
   //Convert the 3rd octet string to numerical value
   STRG_VAL(IN := #tempOctetString,
            FORMAT := W#16#0000,
            P := 1,
            OUT => #tempUInt);
   IF #tempUInt > #MAX_USINT
   THEN
     #error := TRUE;
     #status := #WRONG_VALUE_POS3;
     RETURN;
   ELSE
     #tempIpAdressTaddr.REM_IP_ADDR[3] := UINT_TO_BYTE(#tempUInt);
   END_IF;

   // Process the 4th octet of the IP Address
   #tempCharPosition := FIND(IN1 := #tempAddressString, IN2 := '.');
   IF #tempCharPosition > #NO_POS THEN
     #error := TRUE;
     #status := #WRONG_VALUE_POS4;
     RETURN;
   ELSE
     #tempCharPosition := FIND(IN1 := #tempAddressString, IN2 := ':');
   END_IF;

   // Check if Port number added
   #tempPortNumberIsSpecified := (#tempCharPosition > #NO_POS);
   IF #tempCharPosition > #MAX_CHAR_FOR_PORT_PART THEN
     #error := TRUE;
     #status := #WRONG_VALUE_PORT;
     RETURN;
   END_IF;
   IF NOT #tempPortNumberIsSpecified THEN
     #tempCharPosition := LEN(#tempAddressString) + 1;
   END_IF;

   #tempOctetString := LEFT(IN := #tempAddressString, L := #tempCharPosition - 1);
   // Check if string is empty
   IF #tempOctetString = #EMPTY_STRING THEN
     #error := TRUE;
     #status := #WRONG_VALUE_POS4;
     RETURN;
   ELSE
     #tempAddressString := DELETE(IN := #tempAddressString, P := 1, L := #tempCharPosition);
   END_IF;

   // Convert the 4th octet string to numerical value
   STRG_VAL(IN := #tempOctetString,
            FORMAT := W#16#0000,
            P := 1,
            OUT => #tempUInt);

   IF #tempUInt > #MAX_USINT THEN
     #error := TRUE;
     #status := #WRONG_VALUE_POS4;
     RETURN;
   ELSE
     #tempIpAdressTaddr.REM_IP_ADDR[4] := UINT_TO_BYTE(#tempUInt);
   END_IF;

   // If the string contains a port number too, parse it
   IF #tempPortNumberIsSpecified THEN
     // Convert the port number string to numerical value
     STRG_VAL(IN := #tempAddressString,
              FORMAT := W#16#0000,
              P := 1,
              OUT => #tempUInt);
     IF #tempUInt > #MAX_UINT OR #tempUInt = 0 THEN
       #error := TRUE;
       #status := #WRONG_VALUE_PORT;
       RETURN;
     ELSE
       #tempIpAdressTaddr.REM_PORT_NR := #tempUInt;
     END_IF;
   END_IF;

   // Write Outputs
   #LGF_StringToTaddr := #tempIpAdressTaddr;
END_FUNCTION

ORGANIZATION_BLOCK "Main"   // OB1, LAD, ProgramCycle
TITLE = "Main Program Sweep (Cycle)"
{ S7_Optimized_Access := 'TRUE' }
VERSION : 0.1
   VAR_INPUT
      Initial_Call : Bool;   // Initial call of this OB
      Remanence : Bool;   // =True, if remanent data are available
   END_VAR
   VAR_TEMP
      tmpI : Int;
      tmpI2 : Int;
   END_VAR
BEGIN

REGION Network 2
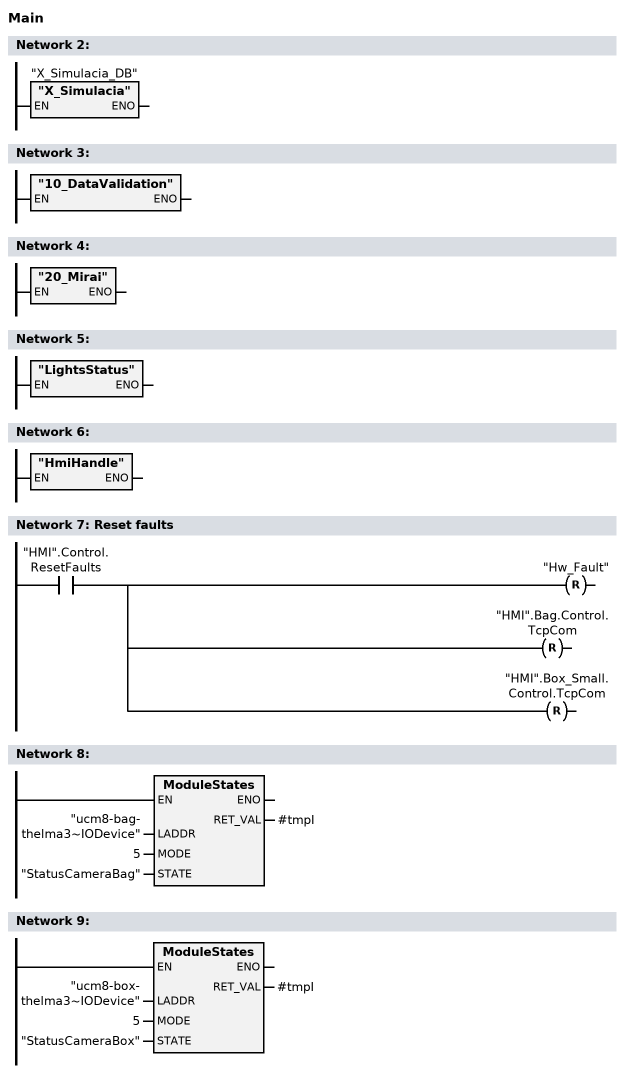
   RUNG wire#powerrail
      "X_Simulacia_DB"()
   END_RUNG
   // the same network as SCL:
   "X_Simulacia_DB"();   // "X_Simulacia"
END_REGION

REGION Network 3
   RUNG wire#powerrail
      "10_DataValidation"()
   END_RUNG
   // the same network as SCL:
   "10_DataValidation"();
END_REGION

REGION Network 4
   RUNG wire#powerrail
      "20_Mirai"()
   END_RUNG
   // the same network as SCL:
   "20_Mirai"();
END_REGION

REGION Network 5
   RUNG wire#powerrail
      "LightsStatus"()
   END_RUNG
   // the same network as SCL:
   "LightsStatus"();
END_REGION

REGION Network 6
   RUNG wire#powerrail
      "HmiHandle"()
   END_RUNG
   // the same network as SCL:
   "HmiHandle"();
END_REGION

REGION Network 7: Reset faults
   RUNG wire#powerrail
      Contact( "HMI".Control.ResetFaults )
      wire#w1
      R_Coil( "Hw_Fault" )
   END_RUNG
   RUNG wire#w1
      R_Coil( "HMI".Bag.Control.TcpCom )
   END_RUNG
   RUNG wire#w1
      R_Coil( "HMI".Box_Small.Control.TcpCom )
   END_RUNG
   // the same network as SCL:
   IF "HMI".Control.ResetFaults THEN
       "Hw_Fault" := FALSE;
       "HMI".Bag.Control.TcpCom := FALSE;
       "HMI".Box_Small.Control.TcpCom := FALSE;
   END_IF;
END_REGION

REGION Network 8
   // no SCL statement known for ModuleStates: written as a call
   #tmpI := ModuleStates(LADDR := "ucm8-bag-thelma3~IODevice", MODE := 5, STATE := "StatusCameraBag");
END_REGION

REGION Network 9
   // no SCL statement known for ModuleStates: written as a call
   #tmpI := ModuleStates(LADDR := "ucm8-box-thelma3~IODevice", MODE := 5, STATE := "StatusCameraBox");
END_REGION
END_ORGANIZATION_BLOCK

ORGANIZATION_BLOCK "Rack or station failure"   // OB86, LAD, RackStationFailure
{ S7_Optimized_Access := 'TRUE' }
VERSION : 0.1
   VAR_INPUT
      LADDR : Hw_Device;   // Hardware identifier
      Event_Class : Byte;   // Event class
      Fault_ID : Byte;   // Fault identifier
   END_VAR
BEGIN

REGION Network 1
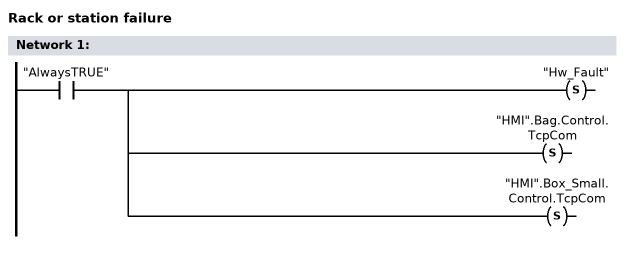
   RUNG wire#powerrail
      Contact( "AlwaysTRUE" )
      wire#w1
      S_Coil( "Hw_Fault" )
   END_RUNG
   RUNG wire#w1
      S_Coil( "HMI".Bag.Control.TcpCom )
   END_RUNG
   RUNG wire#w1
      S_Coil( "HMI".Box_Small.Control.TcpCom )
   END_RUNG
   // the same network as SCL:
   IF "AlwaysTRUE" THEN
       "Hw_Fault" := TRUE;
       "HMI".Bag.Control.TcpCom := TRUE;
       "HMI".Box_Small.Control.TcpCom := TRUE;
   END_IF;
END_REGION
END_ORGANIZATION_BLOCK

ORGANIZATION_BLOCK "Startup"   // OB100, LAD, Startup
TITLE = "Complete Restart"
{ S7_Optimized_Access := 'TRUE' }
VERSION : 0.1
   VAR_INPUT
      LostRetentive : Bool;   // True if retentive data are lost
      LostRTC : Bool;   // True if date and time are lost
   END_VAR
BEGIN

REGION Network 1
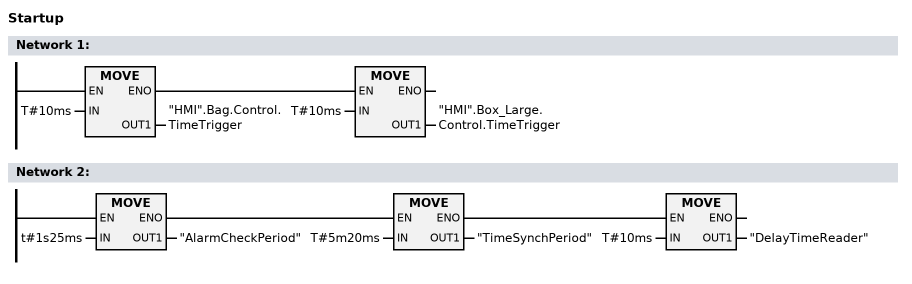
   RUNG wire#powerrail
      Move(in := T#10ms, out1 => "HMI".Bag.Control.TimeTrigger)
      Move(in := T#10ms, out1 => "HMI".Box_Large.Control.TimeTrigger)
   END_RUNG
   // the same network as SCL:
   "HMI".Bag.Control.TimeTrigger := T#10ms;
   "HMI".Box_Large.Control.TimeTrigger := T#10ms;
END_REGION

REGION Network 2
   RUNG wire#powerrail
      Move(in := t#1s25ms, out1 => "AlarmCheckPeriod")
      Move(in := T#5m20ms, out1 => "TimeSynchPeriod")
      Move(in := T#10ms, out1 => "DelayTimeReader")
   END_RUNG
   // the same network as SCL:
   "AlarmCheckPeriod" := t#1s25ms;
   "TimeSynchPeriod" := T#5m20ms;
   "DelayTimeReader" := T#10ms;
END_REGION
END_ORGANIZATION_BLOCK

ORGANIZATION_BLOCK "Programming error"   // OB121, LAD, ProgrammingError
{ S7_Optimized_Access := 'TRUE' }
VERSION : 0.1
   VAR_INPUT
      BlockNr : UInt;   // Number of causing block
      Reaction : USInt;   // 0:ignore, 1:substitute, 2:skip
      Fault_ID : Byte;   // Fault identifier
      BlockType : USInt;   // 16#01:OB, 16#02:FC, 16#03:FB, 16#04:SFC, 16#05:SFB, 16#06:DB: Type of block causing the error
      Area : USInt;   // Area where the error occured
      DBNr : DB_ANY;   // DB number if Area = DB or DI
      Csg_OBNr : OB_Any;   // Number of OB causing the error
      Csg_Prio : USInt;   // Priority of OB causing the error
      Width : USInt;   // 0:bit, 1:byte, 2:word, 3:dword, 4:lword
   END_VAR
BEGIN
END_ORGANIZATION_BLOCK

(* ===== HMI "HMI_RT_2" =====
system functions are stored by id; their names below are inferred from use
connection "HMI_Connection_2": ETHERNET, S7_1500_OMS

HMI tags "Default tag table"
   "screen_titles" : Int, internal
   "system_datetime" : DateTime, internal
   "liuser" : WString[20], internal
   "autoPwd" : WString[10], internal
   "autoUser" : WString[10], internal
   "initDone" : Int, internal

HMI tags "Cam"
   "Rec_HMI_Bag_Cam_Vertiacal_position" : Int = PLC HMI.Bag_Cam.Vertiacal_position, 1 s
   "Rec_HMI_Bag_Cam_Horizontal_position" : Int = PLC HMI.Bag_Cam.Horizontal_position AT %DB1.DBW0, 1 s
   "Rec_HMI_Bag_Cam_Angle" : Int = PLC HMI.Bag_Cam.Angle AT %DB1.DBW0, 1 s
   "Rec_HMI_Box_Cam_Vertiacal_position" : Int = PLC HMI.Box_Cam.Vertiacal_position AT %DB1.DBW0, 1 s
   "Rec_HMI_Box_Cam_Horizontal_position" : Int = PLC HMI.Box_Cam.Horizontal_position AT %DB1.DBW0, 1 s
   "Rec_HMI_Box_Cam_Angle" : Int = PLC HMI.Box_Cam.Angle AT %DB1.DBW0, 1 s
   "Rec_HMI_Bag_Cam_Delay_time_trigger" : Int = PLC HMI.Bag_Cam.Delay_time_trigger AT %DB1.DBW0, 1 s
   "Rec_HMI_Box_Cam_Delay_time_trigger" : Int = PLC HMI.Box_Cam.Delay_time_trigger AT %DB1.DBW0, 1 s
   "SP_HMI_Bag_Cam_Angle" : Int = PLC HMI.Bag_Cam.Angle AT %DB1.DBW0, 1 s
   "SP_HMI_Bag_Cam_Delay_time_trigger" : Int = PLC HMI.Bag_Cam.Delay_time_trigger AT %DB1.DBW0, 1 s
   "SP_HMI_Bag_Cam_Horizontal_position" : Int = PLC HMI.Bag_Cam.Horizontal_position AT %DB1.DBW0, 1 s
   "SP_HMI_Bag_Cam_Vertiacal_position" : Int = PLC HMI.Bag_Cam.Vertiacal_position, 1 s
   "SP_HMI_Box_Cam_Angle" : Int = PLC HMI.Box_Cam.Angle AT %DB1.DBW0, 1 s
   "SP_HMI_Box_Cam_Delay_time_trigger" : Int = PLC HMI.Box_Cam.Delay_time_trigger AT %DB1.DBW0, 1 s
   "SP_HMI_Box_Cam_Horizontal_position" : Int = PLC HMI.Box_Cam.Horizontal_position AT %DB1.DBW0, 1 s
   "SP_HMI_Box_Cam_Vertiacal_position" : Int = PLC HMI.Box_Cam.Vertiacal_position AT %DB1.DBW0, 1 s
   "Rec_HMI_Bag_Cam_Fps" : Int = PLC HMI.Bag_Cam.Fps AT %DB1.DBW0, 1 s
   "Rec_HMI_Box_Cam_Fps" : Int = PLC HMI.Box_Cam.Fps AT %DB1.DBW0, 1 s
   "Rec_HMI_Enigma_off" : Bool = PLC HMI.Enigma_off AT %DB1.DBW0, 1 s
   "Rec_HMI_Mirai_off" : Bool = PLC HMI.Mirai_off AT %DB1.DBX0.0, 1 s
   "SP_HMI_Enigma_off" : Bool = PLC HMI.Enigma_off AT %DB1.DBW0, 1 s
   "SP_HMI_Mirai_off" : Bool = PLC HMI.Mirai_off AT %DB1.DBX0.0, 1 s

HMI tags "Alarms"
   "active_alarms_num" : Int, internal
   "active_alarm" : Bool, internal
   "FaultWord1" : Word = PLC FaultWord1 AT %MW100, 1 s
   "FaultWord2" : Word = PLC FaultWord2 AT %MW102, 1 s
   "FaultWord3" : Word = PLC FaultWord3 AT %MW104, 1 s
   "FaultWord4" : Word = PLC FaultWord4 AT %MW106, 1 s
   "FaultWord5" : Word = PLC FaultWord5 AT %MW108, 1 s
   "FaultWord6" : Word = PLC FaultWord6 AT %MW110, 1 s
   "FaultWord7" : Word = PLC FaultWord7 AT %MW112, 1 s
   "FaultWord8" : Word = PLC FaultWord8 AT %MW114, 1 s

HMI tags "Codes"
   "HMI_Box_Small_Codes_ActualReadingBox" : UDInt = PLC HMI.Box_Small.Codes.ActualReadingBox AT %DB1.DBX0.0, 1 s
   "HMI_Box_Small_Codes_MaterialNumberBox" : UDInt = PLC HMI.Box_Small.Codes.MaterialNumberBox AT %DB1.DBX0.0, 1 s
   "HMI_Bag_Codes_MaterialNumberBox" : UDInt = PLC HMI.Bag.Codes.MaterialNumberBox, 1 s
   "HMI_Bag_Codes_ActualReadingBox" : UDInt = PLC HMI.Bag.Codes.ActualReadingBox, 1 s
   "HMI_Box_Large_Codes_MaterialNumberBox" : String[254] = PLC HMI.Box_Large.Codes.MaterialNumberBox AT %DB1.DBX0.0, 1 s
   "HMI_Box_Large_Codes_ActualReadingBox" : String[254] = PLC HMI.Box_Large.Codes.ActualReadingBox AT %DB1.DBX0.0, 1 s

HMI tags "Control"
   "HMI_Box_Small_Control_ResetCounters" : Bool = PLC HMI.Box_Small.Control.ResetCounters AT %DB1.DBX0.0, 1 s
   "HMI_Bag_Control_ResetCounters" : Bool = PLC HMI.Bag.Control.ResetCounters AT %DB1.DBX0.0, 1 s
   "HMI_Bag_Control_TcpCom" : Bool = PLC HMI.Bag.Control.TcpCom AT %DB1.DBX0.0, 1 s
   "HMI_Box_Small_Control_TcpCom" : Bool = PLC HMI.Box_Small.Control.TcpCom AT %DB1.DBX0.0, 1 s
   "HMI_Box_Small_Control_TimeTrigger" : Time = PLC HMI.Box_Small.Control.TimeTrigger, 1 s
   "HMI_Control_ResetFaults" : Bool = PLC HMI.Control.ResetFaults AT %DB1.DBD0, 1 s
   "HMI_Box_Large_Control_ResetCounters" : Bool = PLC HMI.Box_Large.Control.ResetCounters AT %DB1.DBX0.0, 1 s
   "HMI_Box_Large_Control_TimeTrigger" : Time = PLC HMI.Box_Large.Control.TimeTrigger AT %DB1.DBX0.0, 1 s
   "HMI_Box_Large_Control_TcpCom" : Bool = PLC HMI.Box_Large.Control.TcpCom AT %DB1.DBX0.0, 1 s
   "HMI_Bag_Control_TimeTrigger" : Time = PLC HMI.Bag.Control.TimeTrigger AT %DB1.DBX0.0, 1 s
   "HMI_Control_NewRecipeLoaded" : Bool = PLC HMI.Control.NewRecipeLoaded AT %DB1.DBX0.0, 1 s
   "HMI_Control_AutoRecipeFailed" : Bool = PLC HMI.Control.AutoRecipeFailed AT %DB1.DBX0.0, 1 s

HMI tags "Counters"
   "HMI_Box_Small_Counters_CodeOk" : DInt = PLC HMI.Box_Small.Counters.CodeOk, 1 s
   "HMI_Box_Small_Counters_CodeNok" : DInt = PLC HMI.Box_Small.Counters.CodeNok, 1 s
   "HMI_Box_Small_Counters_CodeBadRead" : DInt = PLC HMI.Box_Small.Counters.CodeBadRead, 1 s
   "HMI_Box_Small_Counters_Trigger" : DInt = PLC HMI.Box_Small.Counters.Trigger, 1 s
   "HMI_Box_Small_Counters_NewData" : DInt = PLC HMI.Box_Small.Counters.NewData, 1 s
   "HMI_Bag_Counters_CodeOk" : DInt = PLC HMI.Bag.Counters.CodeOk AT %DB1.DBD0, 1 s
   "HMI_Bag_Counters_CodeNok" : DInt = PLC HMI.Bag.Counters.CodeNok AT %DB1.DBD0, 1 s
   "HMI_Bag_Counters_CodeBadRead" : DInt = PLC HMI.Bag.Counters.CodeBadRead AT %DB1.DBD0, 1 s
   "HMI_Bag_Counters_Trigger" : DInt = PLC HMI.Bag.Counters.Trigger AT %DB1.DBD0, 1 s
   "HMI_Bag_Counters_NewData" : DInt = PLC HMI.Bag.Counters.NewData AT %DB1.DBD0, 1 s
   "HMI_Box_Small_Counters_NDR" : DInt = PLC HMI.Box_Small.Counters.NDR AT %DB1.DBD0, 1 s
   "HMI_Bag_Counters_NDR" : DInt = PLC HMI.Bag.Counters.NDR AT %DB1.DBD0, 1 s
   "HMI_Box_Large_Counters_CodeOk" : DInt = PLC HMI.Box_Large.Counters.CodeOk AT %DB1.DBD0, 1 s
   "HMI_Box_Large_Counters_CodeNok" : DInt = PLC HMI.Box_Large.Counters.CodeNok AT %DB1.DBD0, 1 s
   "HMI_Box_Large_Counters_CodeBadRead" : DInt = PLC HMI.Box_Large.Counters.CodeBadRead AT %DB1.DBD0, 1 s
   "HMI_Box_Large_Counters_Trigger" : DInt = PLC HMI.Box_Large.Counters.Trigger AT %DB1.DBD0, 1 s
   "HMI_Box_Large_Counters_NewData" : DInt = PLC HMI.Box_Large.Counters.NewData AT %DB1.DBD0, 1 s
   "HMI_Box_Large_Counters_NDR" : DInt = PLC HMI.Box_Large.Counters.NDR AT %DB1.DBD0, 1 s

HMI tags "ActProduction"
   "HMI_line_number_s" : String[254] = PLC HMI.line_number_s, 1 s
   "HMI_order_number_s" : String[254] = PLC HMI.order_number_s, 1 s
   "HMI_article_number_s" : String[254] = PLC HMI.article_number_s, 1 s
   "HMI_product_weight_s" : String[254] = PLC HMI.product_weight_s, 1 s
   "HMI_total_in_bag_s" : String[254] = PLC HMI.total_in_bag_s, 1 s
   "HMI_total_in_box_s" : String[254] = PLC HMI.total_in_box_s, 1 s

HMI tags "MIRAI"
   "AlarmCheckPeriod" : Time = PLC AlarmCheckPeriod AT %MD60, 1 s
   "CON_ConnectHMI" : Bool = PLC CON_ConnectHMI AT %M120.4, 1 s
   "CON_DB_ComandsSending_Video_connected" : Bool = PLC CON_DB.ComandsSending_Video.connected AT %DB1.DBD0, 1 s
   "CON_DB_Domino_ConnectionStatus" : Bool = PLC CON_DB.Domino.ConnectionStatus AT %DB1.DBX0.0, 1 s
   "CON_PrinterConnection" : Bool = PLC CON_PrinterConnection AT %M8.3, 1 s
   "CON_PrinterSelection" : Bool = PLC CON_PrinterSelection AT %M8.0, 1 s
   "DelayTimeReader" : Time = PLC DelayTimeReader AT %MD13, 1 s
   "PrinterData_CON_PrinterBagData_OPC_Error" : Bool = PLC PrinterData.CON.PrinterBagData.OPC_Error AT %DB2.DBX0.0, 1 s
   "OPC_CON_Material_NewBatchEndTime" : String[254] = PLC OPC.CON_Material.NewBatchEndTime AT %DB2.DBX1030.0, 1 s
   "OPC_CON_Material_ActualArtBaseNumber" : String[254] = PLC OPC.CON_Material.ActualArtBaseNumber AT %DB2.DBX1798.0, 1 s
   "OPC_CON_Material_ActualBatchNumber" : String[254] = PLC OPC.CON_Material.ActualBatchNumber AT %DB2.DBX1542.0, 1 s
   "OPC_CON_Material_ActualMarketRegCode" : String[254] = PLC OPC.CON_Material.ActualMarketRegCode AT %DB2.DBX2054.0, 1 s
   "OPC_TRP_Materia_ActualAricleNumber" : String[254] = PLC OPC.TRP_Material.ActualAricleNumber AT %DB2.DBX4108.0, 1 s
   "OPC_TRP_Materia_ActualBatchNumber" : String[254] = PLC OPC.TRP_Material.ActualBatchNumber AT %DB2.DBX3852.0, 1 s
   "OPC_TRP_Materia_ActualGTIN_Number" : String[254] = PLC OPC.TRP_Material.ActualGTIN_Number AT %DB2.DBX3596.0, 1 s
   "PrinterData_CON_PrinterBagData_Date" : String[254] = PLC PrinterData.CON.PrinterBagData.Date AT %DB1.DBX0.0, 1 s
   "PrinterData_CON_PrinterBagData_Initialization" : Bool = PLC PrinterData.CON.PrinterBagData.Initialization AT %DB1.DBX0.0, 1 s
   "PrinterData_CON_PrinterBagData_LED_State" : USInt = PLC PrinterData.CON.PrinterBagData.LED_State AT %DB1.DBX0.0, 1 s
   "PrinterData_CON_PrinterBagData_NonMDR_LabelName" : String[254] = PLC PrinterData.CON.PrinterBagData.NonMDR_LabelName AT %DB1.DBX0.0, 1 s
   "PrinterData_CON_PrinterBagData_RemoteAddress" : String[254] = PLC PrinterData.CON.PrinterBagData.RemoteAddress AT %DB1.DBB0, 1 s
   "PrinterData_CON_PrinterBagData_Time" : String[254] = PLC PrinterData.CON.PrinterBagData.Time AT %DB1.DBX0.0, 1 s
   "PrinterData_TRP_PrinterData_Initialization" : Bool = PLC PrinterData.TRP.PrinterData.Initialization AT %DB1.DBX0.0, 1 s
   "PrinterData_TRP_PrinterData_Inverse" : Bool = PLC PrinterData.TRP.PrinterData.Inverse AT %DB1.DBX0.0, 1 s
   "PrinterData_TRP_PrinterData_LED_State" : USInt = PLC PrinterData.TRP.PrinterData.LED_State AT %DB1.DBX0.0, 1 s
   "PrinterData_TRP_PrinterData_RemoteAddress" : String[254] = PLC PrinterData.TRP.PrinterData.RemoteAddress AT %DB1.DBB0, 1 s
   "PrinterData_TRP_PrinterData_Date" : String[254] = PLC PrinterData.TRP.PrinterData.Date AT %DB1.DBX0.0, 1 s
   "PrinterData_TRP_PrinterData_Time" : String[254] = PLC PrinterData.TRP.PrinterData.Time AT %DB1.DBX0.0, 1 s
   "Reader_TRP_NumGross" : UDInt = PLC Reader.TRP.NumGross AT %DB1.DBB0, 1 s
   "Reader_TRP_NumMisMatch" : UDInt = PLC Reader.TRP.NumMisMatch AT %DB1.DBB0, 1 s
   "Reader_TRP_NumNoRead" : UDInt = PLC Reader.TRP.NumNoRead AT %DB1.DBB0, 1 s
   "Reader_TRP_ResetCounters" : Bool = PLC Reader.TRP.ResetCounters AT %DB1.DBB0, 1 s
   "Reader_TRP_ResetFaults" : Bool = PLC Reader.TRP.ResetFaults AT %DB1.DBB0, 1 s
   "Reader_TRP_MisTriggerFault" : Bool = PLC Reader.TRP.MisTriggerFault AT %DB1.DBX0.0, 1 s
   "TimeSynchPeriod" : Time = PLC TimeSynchPeriod AT %MD64, 1 s
   "TRP_ConnectHMI" : Bool = PLC TRP_ConnectHMI AT %M121.4, 1 s
   "TRP_DB_CommandSending_Markem_connected" : Bool = PLC TRP_DB.CommandSending_Markem.connected AT %DB1.DBB0, 1 s
   "TRP_DB_MarkemImaje_ConnectionStatus" : Bool = PLC TRP_DB.MarkemImaje.ConnectionStatus AT %DB1.DBB0, 1 s
   "TRP_DB_MarkemImaje_ExtDate" : String[254] = PLC TRP_DB.MarkemImaje.ExtDate AT %DB1.DBX0.0, 1 s
   "OPC_CON_Material_BatchStatus" : Byte = PLC OPC.CON_Material.BatchStatus, 1 s
   "OPC_CON_Material_NewMarketREG_Code" : String[254] = PLC OPC.CON_Material.NewMarketREG_Code AT %DB1.DBX0.0, 1 s
   "OPC_TRP_Materia_NewGTIN_Number" : String[254] = PLC OPC.TRP_Material.NewGTIN_Number AT %DB1.DBX0.0, 1 s
   "CON_DB_HandleComBag_ActualArtFlag" : Bool = PLC CON_DB.HandleComBag.ActualArtFlag, 1 s
   "CON_DB_HandleComBag_ActualMDR_Flag" : Bool = PLC CON_DB.HandleComBag.ActualMDR_Flag, 1 s
   "OPC_CON_Material_ActualBBD" : String[254] = PLC OPC.CON_Material.ActualBBD, 1 s
   "OPC_CON_Material_NewArtBaseNumber" : UDInt = PLC OPC.CON_Material.NewArtBaseNumber, 1 s
   "OPC_CON_Material_NewArticleFlag" : String[254] = PLC OPC.CON_Material.NewArticleFlag, 1 s
   "OPC_CON_Material_NewBatchNumber" : String[254] = PLC OPC.CON_Material.NewBatchNumber, 1 s
   "OPC_CON_Material_NewBBD" : String[254] = PLC OPC.CON_Material.NewBBD, 1 s
   "OPC_CON_Material_NewMDR_Flag" : String[254] = PLC OPC.CON_Material.NewMDR_Flag, 1 s
   "OPC_TRP_Materia_ActualMachineID" : String[254] = PLC OPC.TRP_Material.ActualMachineID, 1 s
   "OPC_TRP_Materia_NewArticleNumber" : UDInt = PLC OPC.TRP_Material.NewArticleNumber, 1 s
   "OPC_TRP_Materia_NewMachineID" : String[254] = PLC OPC.TRP_Material.NewMachineID, 1 s
   "PrinterData_CON_PrinterSelection" : Bool = PLC PrinterData.CON.PrinterSelection, 1 s
   "Reader_TRP_NumMatch" : UDInt = PLC Reader.TRP.NumMatch, 1 s
   "TRP_DB_MarkemImaje_ExpFlag" : Bool = PLC TRP_DB.MarkemImaje.ExpFlag, 1 s
   "TRP_DB_MarkemImaje_Serial" : UDInt = PLC TRP_DB.MarkemImaje.Serial, 1 s
   "TRP_DB_MarkemImaje_TimePrinted" : String[254] = PLC TRP_DB.MarkemImaje.TimePrinted, 1 s
   "TRP_DB_Reader_2D_Instance_TriggerReady" : Bool = PLC TRP_DB.Reader_2D_Instance.TriggerReady AT %DB1.DBX0.0, 1 s

HMI tags "Recipe"
   "Rec_DeleteResult" : Int, internal
   "Rec_EditResult" : Int, internal
   "Rec_FunctionResultSwitch" : Int, internal
   "Rec_FunctionUsed" : Int, internal
   "Rec_LoadResult" : Int, internal
   "Rec_ReadSPResult" : Int, internal
   "Rec_SaveResult" : Int, internal
   "Rec_SelectedRecipe" : WString[50], internal
   "Rec_ViewResult" : Int, internal
   "INT_0" : Int, internal
   "Rec_AutoSelectResult" : Int = PLC HMI.Control.Status AT %DB1.DBW0, 1 s
   "PlainHandle_DB_NewArticleNum" : String[254] = PLC PlainHandle_DB.NewArticleNum, 1 s
   "FindRecipe" : Bool = PLC FindRecipe AT %M18.1, 1 s
      on ChangeValue: "Rec_AutoSelectRecipe"()

HMI tags "Service"
   "X_Simulacia_DB_TRP_Materia_NewGTIN_Number" : String[254] = PLC X_Simulacia_DB.TRP_Materia.NewGTIN_Number, 1 s
   "X_Simulacia_DB_TRP_Materia_NewBatchNumber" : String[254] = PLC X_Simulacia_DB.TRP_Materia.NewBatchNumber, 1 s
   "X_Simulacia_DB_TRP_Materia_NewArticleNumber" : UDInt = PLC X_Simulacia_DB.TRP_Materia.NewArticleNumber, 1 s
   "X_Simulacia_DB_TRP_Materia_NewMachineID" : String[254] = PLC X_Simulacia_DB.TRP_Materia.NewMachineID, 1 s
   "X_Simulacia_DB_TRP_Materia_NewBBD" : String[254] = PLC X_Simulacia_DB.TRP_Materia.NewBBD, 1 s
   "X_Simulacia_DB_BagServis" : String[254] = PLC X_Simulacia_DB.BagServis AT %DB1.DBX0.0, 1 s
   "X_Simulacia_DB_BoxServis" : String[254] = PLC X_Simulacia_DB.BoxServis AT %DB1.DBX0.0, 1 s
   "X_Simulacia_DB_Servis_Bag" : Bool = PLC X_Simulacia_DB.Servis.Bag AT %DB1.DBX0.0, 1 s
   "X_Simulacia_DB_Servis_BoxSmall" : Bool = PLC X_Simulacia_DB.Servis.BoxSmall AT %DB1.DBX0.0, 1 s
   "X_Simulacia_DB_Servis_BoxLarge" : Bool = PLC X_Simulacia_DB.Servis.BoxLarge AT %DB1.DBX0.0, 1 s

discrete alarms
   1: 'VIDEOJET/DOMINO chybná IP / VIDEOJET/DOMINO Error IP', class Warnings, trigger "FaultWord1" bit 8
   2: 'VIDEOJET/DOMINO chyba komunikácie / VIDEOJET/DOMINO communication error', class Warnings, trigger "FaultWord1" bit 9
   3: 'A_F1_2', class Warnings, trigger "FaultWord1" bit 10
   4: 'A_F1_3', class Warnings, trigger "FaultWord1" bit 11
   5: 'Žiadne dáta z Plainu / No data from plain', class Warnings, trigger "FaultWord1" bit 12
   6: 'Chyba komunikácie Plain / Communication error plain', class Warnings, trigger "FaultWord1" bit 13
   7: 'Žiadne nové dáta z Plainu / No new data from plain', class Warnings, trigger "FaultWord1" bit 14
   8: 'A_F1_7', class Warnings, trigger "FaultWord1" bit 15
   9: 'Prístup IO prerušený / Access IO disrupted', class Warnings, trigger "FaultWord1" bit 0
   10: 'BOX 3 po sebe nezhodné / BOX 3 not matching in row', class Warnings, trigger "FaultWord1" bit 1
   11: 'BOX 3 po sebe nezhodné/neprečítané / BOX 3 no readings in a row', class Warnings, trigger "FaultWord1" bit 2
   12: 'Chyba senzor BOX / BOX trigger not ready', class Warnings, trigger "FaultWord1" bit 3
   13: 'Enigma zakázaná / Disable Enigma', class Warnings, trigger "FaultWord1" bit 4
   14: 'Neplatné číslo materiálu pre BOX / Not valid material number for box', class Warnings, trigger "FaultWord1" bit 5
   15: 'A_F1_14', class Warnings, trigger "FaultWord1" bit 6
   16: 'A_F1_15', class Warnings, trigger "FaultWord1" bit 7
   17: 'Platnosť Batch sa blíži ku koncu / Batch end time warning', class Warnings, trigger "FaultWord2" bit 8
   18: 'Platnosť Batch vypršala / Batch end time error', class Warnings, trigger "FaultWord2" bit 9
   19: 'A_F2_2', class Warnings, trigger "FaultWord2" bit 10
   20: 'A_F2_3', class Warnings, trigger "FaultWord2" bit 11
   21: 'A_F2_4', class Warnings, trigger "FaultWord2" bit 12
   22: 'A_F2_5', class Warnings, trigger "FaultWord2" bit 13
   23: 'A_F2_6', class Warnings, trigger "FaultWord2" bit 14
   24: 'A_F2_7', class Warnings, trigger "FaultWord2" bit 15
   25: 'A_F2_8', class Warnings, trigger "FaultWord2" bit 0
   26: 'BAG 3 po sebe nezhodné / BAG 3 not matching in row', class Warnings, trigger "FaultWord2" bit 1
   27: 'BAG 3 po sebe neprečítané / BAG 3 no reading in a row', class Warnings, trigger "FaultWord2" bit 2
   28: 'Chyba senzor BAG / BAG trigger watchdog', class Warnings, trigger "FaultWord2" bit 3
   29: 'Enigma zakázaná pre BAG / Enigma Disable for BAG', class Warnings, trigger "FaultWord2" bit 4
   30: 'Neplatné číslo materiálu pre BAG / Not valid material number for BAG', class Warnings, trigger "FaultWord2" bit 5
   31: 'A_F2_14', class Warnings, trigger "FaultWord2" bit 6
   32: 'A_F2_15', class Warnings, trigger "FaultWord2" bit 7
   33: 'A_F6_0', class Warnings, trigger "FaultWord6" bit 8
   34: 'A_F6_1', class Warnings, trigger "FaultWord6" bit 9
   35: 'A_F6_2', class Warnings, trigger "FaultWord6" bit 10
   36: 'A_F6_3', class Warnings, trigger "FaultWord6" bit 11
   37: 'A_F6_4', class Warnings, trigger "FaultWord6" bit 12
   38: 'HW chyba / HW Faults', class Warnings, trigger "FaultWord6" bit 13
   39: 'A_F6_6', class Warnings, trigger "FaultWord6" bit 14
   40: 'A_F6_7', class Warnings, trigger "FaultWord6" bit 15
   41: 'Chyba kamera BAG / Fault reader BAG', class Warnings, trigger "FaultWord6" bit 0
   42: 'Chyba kamera BOX / Fault reader BOX', class Warnings, trigger "FaultWord6" bit 1
   43: 'BOX kamera zle prečítala / BOX Reader had no good reading', class Warnings, trigger "FaultWord6" bit 2
   44: 'A_F6_11', class Warnings, trigger "FaultWord6" bit 3
   45: 'A_F6_12', class Warnings, trigger "FaultWord6" bit 4
   46: 'A_F6_13', class Warnings, trigger "FaultWord6" bit 5
   47: 'A_F6_14', class Warnings, trigger "FaultWord6" bit 6
   48: 'A_F6_15', class Warnings, trigger "FaultWord6" bit 7
   49: 'A_F7_0', class Warnings, trigger "FaultWord7" bit 8
   50: 'A_F7_1', class Warnings, trigger "FaultWord7" bit 9
   51: 'BAG kamera zle prečítala / BAG Reader had no good reading', class Warnings, trigger "FaultWord7" bit 10
   52: 'A_F7_3', class Warnings, trigger "FaultWord7" bit 11
   53: 'A_F7_4', class Warnings, trigger "FaultWord7" bit 12
   54: 'A_F7_5', class Warnings, trigger "FaultWord7" bit 13
   55: 'A_F7_6', class Warnings, trigger "FaultWord7" bit 14
   56: 'A_F7_7', class Warnings, trigger "FaultWord7" bit 15
   57: 'A_F7_8', class Warnings, trigger "FaultWord7" bit 0
   58: 'A_F7_9', class Warnings, trigger "FaultWord7" bit 1
   59: 'A_F7_10', class Warnings, trigger "FaultWord7" bit 2
   60: 'A_F7_11', class Warnings, trigger "FaultWord7" bit 3
   61: 'A_F7_12', class Warnings, trigger "FaultWord7" bit 4
   62: 'A_F7_13', class Warnings, trigger "FaultWord7" bit 5
   63: 'A_F7_14', class Warnings, trigger "FaultWord7" bit 6
   64: 'A_F7_15', class Warnings, trigger "FaultWord7" bit 7
   65: 'A_F3_0', class Warnings, trigger "FaultWord3" bit 8
   67: 'A_F3_2', class Warnings, trigger "FaultWord3" bit 10
   68: 'A_F3_3', class Warnings, trigger "FaultWord3" bit 11
   69: 'A_F3_4', class Warnings, trigger "FaultWord3" bit 12
   70: 'A_F3_5', class Warnings, trigger "FaultWord3" bit 13
   71: 'A_F3_6', class Warnings, trigger "FaultWord3" bit 14
   72: 'A_F3_7', class Warnings, trigger "FaultWord3" bit 15
   73: 'TRP chybná IP / TRP Error IP', class Warnings, trigger "FaultWord3" bit 0
   74: 'TRP chyba komunikácie / TRP Communication error', class Warnings, trigger "FaultWord3" bit 1
   75: 'A_F3_10', class Warnings, trigger "FaultWord3" bit 2
   76: 'A_F3_11', class Warnings, trigger "FaultWord3" bit 3
   77: 'A_F3_12', class Warnings, trigger "FaultWord3" bit 4
   78: 'A_F3_13', class Warnings, trigger "FaultWord3" bit 5
   79: 'A_F3_14', class Warnings, trigger "FaultWord3" bit 6
   80: 'A_F3_15', class Warnings, trigger "FaultWord3" bit 7
   81: 'Label print istič chyba -01FA6 / Label print breaker error -01FA6', class Warnings, trigger "FaultWord4" bit 8
   82: 'Napajanie DI istič chyba -03FA5 / Power source DI breaker error -03FA5', class Warnings, trigger "FaultWord4" bit 9
   83: 'Napájanie Ventilátor chyba -03FA6 / Power source fan breaker error -03FA6', class Warnings, trigger "FaultWord4" bit 10
   84: 'A_F4_3', class Warnings, trigger "FaultWord4" bit 11
   85: 'A_F4_4', class Warnings, trigger "FaultWord4" bit 12
   86: 'A_F4_5', class Warnings, trigger "FaultWord4" bit 13
   87: 'A_F4_6', class Warnings, trigger "FaultWord4" bit 14
   88: 'A_F4_7', class Warnings, trigger "FaultWord4" bit 15
   89: 'MIRAI 3 po sebe neprečítané / MIRAI 3 not reading in row', class Warnings, trigger "FaultWord4" bit 0
   90: 'MIRAI 3 po sebe nezhodné / MIRAI 3 not matching in row', class Warnings, trigger "FaultWord4" bit 1
   91: 'A_F4_10', class Warnings, trigger "FaultWord4" bit 2
   92: 'A_F4_11', class Warnings, trigger "FaultWord4" bit 3
   93: 'A_F4_12', class Warnings, trigger "FaultWord4" bit 4
   94: 'A_F4_13', class Warnings, trigger "FaultWord4" bit 5
   95: 'A_F4_14', class Warnings, trigger "FaultWord4" bit 6
   96: 'A_F4_15', class Warnings, trigger "FaultWord4" bit 7
   97: 'TRP Printer Fault/Warning: / TRP tlačiareň Chyba/Varovanie', class Warnings, trigger "FaultWord5" bit 8
   98: 'TRP Printer Fault/Warning: / TRP tlačiareň Chyba/Varovanie', class Warnings, trigger "FaultWord5" bit 9
   99: 'TRP Printer Fault/Warning: / TRP tlačiareň Chyba/Varovanie', class Warnings, trigger "FaultWord5" bit 10
   100: 'TRP Printer Fault/Warning: / TRP tlačiareň Chyba/Varovanie', class Warnings, trigger "FaultWord5" bit 11
   101: 'TRP Printer Fault/Warning: / TRP tlačiareň Chyba/Varovanie', class Warnings, trigger "FaultWord5" bit 12
   102: 'TRP Printer Fault/Warning: / TRP tlačiareň Chyba/Varovanie', class Warnings, trigger "FaultWord5" bit 13
   103: 'TRP Printer Fault/Warning: / TRP tlačiareň Chyba/Varovanie', class Warnings, trigger "FaultWord5" bit 14
   104: 'TRP Printer Fault/Warning: / TRP tlačiareň Chyba/Varovanie', class Warnings, trigger "FaultWord5" bit 15
   105: 'TRP Printer Fault/Warning: / TRP tlačiareň Chyba/Varovanie', class Warnings, trigger "FaultWord5" bit 0
   106: 'TRP Printer Fault/Warning: / TRP tlačiareň Chyba/Varovanie', class Warnings, trigger "FaultWord5" bit 1
   107: 'TRP Printer Fault/Warning: / TRP tlačiareň Chyba/Varovanie', class Warnings, trigger "FaultWord5" bit 2
   108: 'TRP Printer Fault/Warning: / TRP tlačiareň Chyba/Varovanie', class Warnings, trigger "FaultWord5" bit 3
   109: 'TRP Printer Fault/Warning: / TRP tlačiareň Chyba/Varovanie', class Warnings, trigger "FaultWord5" bit 4
   110: 'TRP Printer Fault/Warning: / TRP tlačiareň Chyba/Varovanie', class Warnings, trigger "FaultWord5" bit 5
   111: 'TRP Printer Fault/Warning: / TRP tlačiareň Chyba/Varovanie', class Warnings, trigger "FaultWord5" bit 6
   112: 'TRP Printer Fault/Warning: / TRP tlačiareň Chyba/Varovanie', class Warnings, trigger "FaultWord5" bit 7
   66: 'A_F3_1', class Warnings, trigger "FaultWord3" bit 9
   113: 'TRP Printer Fault/Warning: / TRP tlačiareň Chyba/Varovanie', class Warnings, trigger "FaultWord8" bit 8
   114: 'TRP Printer Fault/Warning: / TRP tlačiareň Chyba/Varovanie', class Warnings, trigger "FaultWord8" bit 9
   115: 'TRP Printer Fault/Warning: / TRP tlačiareň Chyba/Varovanie', class Warnings, trigger "FaultWord8" bit 10
   116: 'TRP Printer Fault/Warning: / TRP tlačiareň Chyba/Varovanie', class Warnings, trigger "FaultWord8" bit 11
   117: 'TRP Printer Fault/Warning: / TRP tlačiareň Chyba/Varovanie', class Warnings, trigger "FaultWord8" bit 12
   118: 'TRP Printer Fault/Warning: / TRP tlačiareň Chyba/Varovanie', class Warnings, trigger "FaultWord8" bit 13
   119: 'TRP Printer Fault/Warning: / TRP tlačiareň Chyba/Varovanie', class Warnings, trigger "FaultWord8" bit 14
   120: 'TRP Printer Fault/Warning: / TRP tlačiareň Chyba/Varovanie', class Warnings, trigger "FaultWord8" bit 15
   121: 'TRP Printer Fault/Warning: / TRP tlačiareň Chyba/Varovanie', class Warnings, trigger "FaultWord8" bit 0
   122: 'TRP Printer Fault/Warning: / TRP tlačiareň Chyba/Varovanie', class Warnings, trigger "FaultWord8" bit 1
   123: 'TRP Printer Fault/Warning: / TRP tlačiareň Chyba/Varovanie', class Warnings, trigger "FaultWord8" bit 2
   124: 'TRP Printer Fault/Warning: / TRP tlačiareň Chyba/Varovanie', class Warnings, trigger "FaultWord8" bit 3
   125: 'TRP Printer Fault/Warning: / TRP tlačiareň Chyba/Varovanie', class Warnings, trigger "FaultWord8" bit 4
   126: 'TRP Printer Fault/Warning: / TRP tlačiareň Chyba/Varovanie', class Warnings, trigger "FaultWord8" bit 5
   127: 'TRP Printer Fault/Warning: / TRP tlačiareň Chyba/Varovanie', class Warnings, trigger "FaultWord8" bit 6
   128: 'TRP Printer Fault/Warning:/Warning:/Warning: / TRP tlačiareň Chyba/Varovanie', class Warnings, trigger "FaultWord8" bit 7

text list "CON_Printers": 0 'Domino'; 1 'Video Jet'

text list "screenTitle": 1 'ENIGMA Overview ENIGMA Prehľad'; 2 'Alarms / História alarmov'; 7 'ENIGMA Settings - trigger delay ENIGMA Nastavenia - oneskorenie čítania'; 8 'ENIGMA Settings - camera position ENIGMA Nastavania - pozícia kamery'; 3 'ENIGMA Status'; 20 'System / Systém'; 23 'System - user administration / Správa používateľov'; 4 'Recipe selection / Výber receptu'; 0 'Package validation / Validácia balení'; 5 'Recipe viewer / Prehliadač receptov'; 6 'Recipe editor / Editor receptov'; 25 'System - diagnostics / Diagnostika systému'; 50 'MIRAI Overview MIRAI Prehľad'; 52 'MIRAI Settings - printer MIRAI Nastavenia - tlačiaren'; 51 'MIRAI Status'; 53 'MIRAI Settings - trigger delay MIRAI Nastavenia - oneskorenie čítania'; 60 'Service / Servis'; 26 'Systémové nastavenia / System settings'; 24 'Iné nástroje / Other tools'; 21 'Informácie o projekte / Project information'; 22 'Informácie o systéme / System information'; 54 'MIRAI Settings - camera position MIRAI Nastavenia - pozícia kamery'

text list "TRP_PrinterErrorsW1": 8 'Overheated / Systém je prehriaty'; 9 'I/O board error / Chyba vstupno/výstupnej dosky'; 10 'File system error / Chyba súborov'; 11 'Memory error / Chyba pamäte'; 12 'Parameter error / Chyba parametrov'; 13 'No init file / Inicializačný súbor nie je prítomný'; 14 'No air pressure / Chyba tlaku vzduchu'; 15 'Paper out / Papier neprítomný'; 0 'Ribbon out / Páska minutá'; 1 'Head lifted / Hlava je zdvihnutá'; 2 'Press start / Stlač štart'; 3 'No return signal / Žiadna spätná väzba'; 4 'Arm jammed / Nanášacia hlavica zaseknutá'; 5 'Arm not home / Nanášacia hlavica nie je v základnej polohe'; 6 'Barcode error / Chyba barkódu'; 7 'Label on grid / Štíkok je na mriežke'

text list "TRP_PrinterErrorsW2": 8 'No label on grid / Žiadny štíkok na hlavici'; 9 'Cover open / Kryt otvorený'; 10 'Pause / Pauza'; 11 'Paper low / Dochádza papier'; 12 'Ribbon low / Dochádza kotúč'; 13 'Barcode warning / Varovanie barkód'; 14 'ApplyDelay too short / Oneskorenie nanášania je príliš nízke'; 15 'Accept date change / Prijať zmenu údajov'; 0 'Matchcode error / Chyba zhody kódu'; 1 'Barcode quality / Chyba kvality barkódu'; 2 'Waiting for trig / Čakám na spúšťací signál'; 3 'Trig Sensor Error / Chyba trigrovacieho senzoru'; 4 'Printer Synchronization / Synchronizácia tlačiarne'; 5 'Printer Synchronization Timeout / Čas pre synchronizáciu tlačiarne vypršal'; 6 'Product Too Close / Produkt je príliš blízko'; 7 'SSCC limit reached / SSCC limit dosiahnutý'

graphic list "On_Off_NonEditable": 0 'checkbox_checked_disabled'; 1 'checkbox_empty_disabled'

graphic list "On_Off_Editable": 0 'checkbox_checked'; 1 'checkbox_empty'

recipe "ReaderRecipes": bag_horizontal_pos <- "Rec_HMI_Bag_Cam_Horizontal_position", bag_vertical_pos <- "Rec_HMI_Bag_Cam_Vertiacal_position", bag_angle <- "Rec_HMI_Bag_Cam_Angle", bag_trigger_delay <- "Rec_HMI_Bag_Cam_Delay_time_trigger", box_horizontal_pos <- "Rec_HMI_Box_Cam_Horizontal_position", box_vertical_pos <- "Rec_HMI_Box_Cam_Vertiacal_position", box_angle <- "Rec_HMI_Box_Cam_Angle", box_trigger_delay <- "Rec_HMI_Box_Cam_Delay_time_trigger", bag_fps <- "Rec_HMI_Bag_Cam_Fps", box_fps <- "Rec_HMI_Box_Cam_Fps", enima_off <- "Rec_HMI_Enigma_off", mirai_off <- "Rec_HMI_Mirai_off"

screen "Menu" 800x414
   on GenerateScreen: SetTag("screen_titles", 0)
   Button "Button_1" at 333,16 size 135x52; TextOff 'Enigma'
      on Release: ActivateScreen("MainScreen", 0)
   Button "Button_2" at 333,88 size 135x52; TextOff 'Mirai'
      on Release: ActivateScreen("Main", 0)
   Button "Button_3" at 333,160 size 135x52; TextOff 'Service / Servis'; Authorization "User administration"
      on Release: ActivateScreen("Service", 0)
   Button "Button_4" at 513,232 size 135x90; TextOff 'Enigma'; PictureOff "Slovakia"
      on Click: function_fb9197e8(L sk-SK)
   Button "Button_5" at 657,232 size 135x90; TextOff 'Enigma'; PictureOff "United_Kingdom"
      on Click: function_fb9197e8(L en-US)

screen "Main" 800x414, template "Template_Mirai"
   on GenerateScreen: SetTag("screen_titles", 50)
   TextField "Text field_1" at 497,27 size 301x23; Text 'Camera / Kamera'
   TextField "Text field_2" at 274,4 size 212x32; Text 'Batch End Time / Koniec objednávky'
   TextField "Text field_3" at 520,61 size 107x23; Text '# Triggers / # Zosnímané'
   TextField "Text field_4" at 520,95 size 111x23; Text '# No-Reads / # Neprečítané'
   TextField "Text field_5" at 520,131 size 113x23; Text '# Mis-Match / # Nezhodné'
   IOField "I/O field_1" at 632,61 size 148x23; FormatPattern 9999999999
      ProcessValue <- "Reader_TRP_NumGross"
   IOField "I/O field_2" at 632,95 size 148x23; FormatPattern 9999999999
      ProcessValue <- "Reader_TRP_NumNoRead"
   IOField "I/O field_3" at 632,131 size 148x23; FormatPattern 9999999999
      ProcessValue <- "Reader_TRP_NumMisMatch"
   IOField "I/O field_4" at 291,56 size 177x32; FormatPattern ????????????????????
      ProcessValue <- "OPC_CON_Material_NewBatchEndTime"
   Circle "Circle_1" at 470,55 size 34x34
      Appearance <- "OPC_CON_Material_BatchStatus"
   TextField "Text field_6" at 16,60 size 120x23; Text 'TRP Printer / TRP tlačiareň'
   TextField "Text field_7" at 16,100 size 120x23; Text 'CON Printer / CON tlačiareň'
   TextField "Text field_8" at 16,140 size 107x23; Text 'Plain'
   TextField "Text field_9" at 16,180 size 107x23; Text 'Reader / Kamera'
   TextField "Text field_10" at 16,220 size 107x23; Text 'Trigger / Senzor'
   Circle "Circle_2" at 136,55 size 34x34
      Appearance <- "TRP_DB_MarkemImaje_ConnectionStatus"
   Circle "Circle_3" at 205,55 size 34x34
      Appearance <- "PrinterData_TRP_PrinterData_LED_State"
   Circle "Circle_4" at 136,95 size 34x34
      Appearance <- "CON_PrinterConnection"
   Circle "Circle_6" at 136,135 size 34x34
      Appearance <- "PrinterData_CON_PrinterBagData_OPC_Error"
   Circle "Circle_9" at 205,175 size 34x34
      Appearance <- "TRP_DB_Reader_2D_Instance_TriggerReady"
   Circle "Circle_11" at 205,215 size 34x34
      Appearance <- "Reader_TRP_MisTriggerFault"
   TextField "Text field_11" at 94,27 size 108x23; Text 'Connection / Spojenie'
   TextField "Text field_12" at 197,27 size 66x23; Text 'Status'
   Button "Button_1" at 676,220 size 104x32; TextOff 'RESET'
      on Release: ResetBit("HMI_Box_Large_Control_ResetCounters")
      on Press: SetBit("HMI_Box_Large_Control_ResetCounters")
   TextField "Text field_13" at 520,169 size 113x23; Text '# Match / # Zhodné'
   IOField "I/O field_5" at 632,169 size 148x23; FormatPattern 9999999999
      ProcessValue <- "Reader_TRP_NumMatch"
   Circle "Circle_7" at 205,95 size 34x34
      Appearance <- "PrinterData_CON_PrinterBagData_LED_State"
   SymbolicIOField "Symbolic I/O field_1" at 291,102 size 175x32; TextOff 'Normal Products / Normal Produkt'; TextOn 'Medical Products / Medical Produkt'
      ProcessValue <- "CON_DB_HandleComBag_ActualMDR_Flag"

